(* Logix 5000 project; controller FV vendor 1 type 14 code 217 rev 31.11; software revision 31.00; part 14 of 63 *)
(* tags used below, declared in another part *)
   CWD : CHECKWORD_FLAGS;
   FR_B240 : INT[255];   // DEBOUNCE Debounce Flags
   FR_B246 : INT[255];   // V_REVERSE Flags for reversing contol action
   FR_B3 : INT[255];   // BINARY
   FR_data_file_value_to_move : DINT;
   FR_F102 : REAL[20];
   FR_FV31_AV01 : PlantItem;   // FV31_AV01
   FR_FV31_AV04 : PlantItem;   // FV31_AV04
   FR_FV31_AV05 : PlantItem;   // FV31_AV05
   FR_FV31_AV06 : PlantItem;   // FV31_AV06
   FR_FV31_AV07 : PlantItem;   // FV31_AV07
   FR_FV31_ROTO : PlantItem;   // FV31_ROTO
   FR_FV31_VA01 : PlantItem;   // FV31_VA01
   FR_N10 : INT[265];   // FV_AGING Comms to FV Aging PL C
   FR_N100 : INT[265];   // FV FILLING
   FR_N110 : INT[265];   // GREEN BEER Green Beer Main
   FR_N120 : INT[265];   // YEAST CROP Yeast Cropping Main
   FR_N13 : INT[265];   // MV_ROUTE Comms to MV Routing PLC
   FR_N130 : INT[265];   // FILTRATE Filtrate Return
   FR_N14 : INT[265];   // MVFV CIP Comms to MVFV CIP Un it PLC
   FR_N160 : INT[265];   // VESSEL Vessel Working Direc tory
   FR_N200 : INT[265];   // ANALOG_IN Analog Inputs
   FR_N255 : INT[265];   // CHECKWORDS
   FR_N31 : INT[265];   // FV31
   FR_N7 : INT[265];   // INTEGER
   FR_N99 : INT[265];   // COMMENT Comment Lines
   FR_OXY_SW1 : PlantItem;   // OXY_SW1
   FR_OXY_SW2 : PlantItem;   // OXY_SW2
   FR_T101 : TIMER[255];   // FV FILLING
   FR_T144 : TIMER[255];   // CIP
   FR_T4 : TIMER[255];   // TIMER
   FR_T50 : TIMER[52];
   FR_T51 : TIMER[52];
   FR_T52 : TIMER[52];
   FR_T53 : TIMER[52];
   FR_VB1_AV08 : PlantItem;   // VB1_AV08
   FR_VB1_AV09 : PlantItem;   // VB1_AV09
   FR_VB2_AV04 : PlantItem;   // VB2_AV04
   FR_VB2_AV05 : PlantItem;   // VB2_AV05
   FR_VB3_AV04 : PlantItem;   // VB3_AV04
   FR_VB3_AV05 : PlantItem;   // VB3_AV05
   FR_VB4_AV03 : PlantItem;   // VB4_AV03
   FR_VB4_AV09 : PlantItem;   // VB4_AV09
   FR_VB4_AV15 : PlantItem;   // VB4_AV15
(* FR_Common, continued *)

ROUTINE FR_FV31_31   (* ladder *)
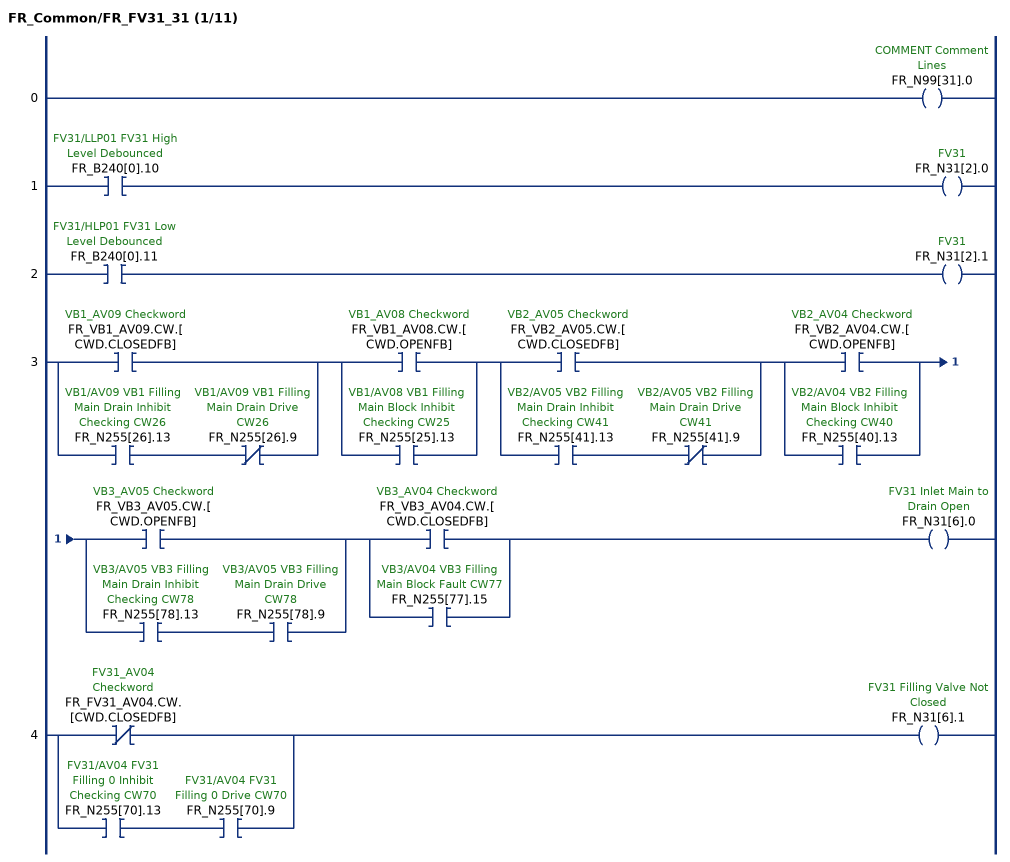
   0: OTE(FR_N99[31].0);
   1: XIC(FR_B240[0].10)OTE(FR_N31[2].0);
   2: XIC(FR_B240[0].11)OTE(FR_N31[2].1);
   3: [XIC(FR_VB1_AV09.CW.[CWD.CLOSEDFB]) ,XIC(FR_N255[26].13) XIO(FR_N255[26].9) ][XIC(FR_VB1_AV08.CW.[CWD.OPENFB]) ,XIC(FR_N255[25].13) ][XIC(FR_VB2_AV05.CW.[CWD.CLOSEDFB]) ,XIC(FR_N255[41].13) XIO(FR_N255[41].9) ][XIC(FR_VB2_AV04.CW.[CWD.OPENFB]) ,XIC(FR_N255[40].13) ][XIC(FR_VB3_AV05.CW.[CWD.OPENFB]) ,XIC(FR_N255[78].13) XIC(FR_N255[78].9) ][XIC(FR_VB3_AV04.CW.[CWD.CLOSEDFB]) ,XIC(FR_N255[77].15) ]OTE(FR_N31[6].0);
   4: [XIO(FR_FV31_AV04.CW.[CWD.CLOSEDFB]) ,XIC(FR_N255[70].13) XIC(FR_N255[70].9) ]OTE(FR_N31[6].1);
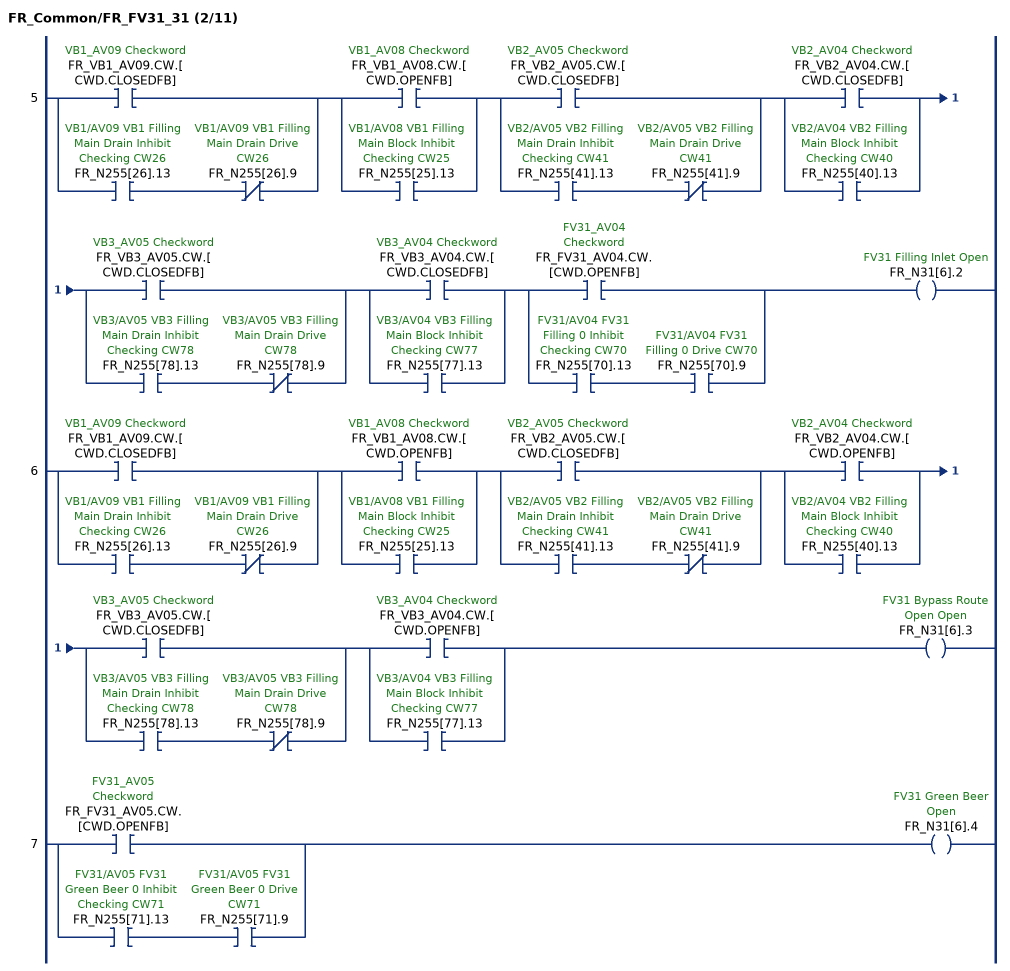
   5: [XIC(FR_VB1_AV09.CW.[CWD.CLOSEDFB]) ,XIC(FR_N255[26].13) XIO(FR_N255[26].9) ][XIC(FR_VB1_AV08.CW.[CWD.OPENFB]) ,XIC(FR_N255[25].13) ][XIC(FR_VB2_AV05.CW.[CWD.CLOSEDFB]) ,XIC(FR_N255[41].13) XIO(FR_N255[41].9) ][XIC(FR_VB2_AV04.CW.[CWD.CLOSEDFB]) ,XIC(FR_N255[40].13) ][XIC(FR_VB3_AV05.CW.[CWD.CLOSEDFB]) ,XIC(FR_N255[78].13) XIO(FR_N255[78].9) ][XIC(FR_VB3_AV04.CW.[CWD.CLOSEDFB]) ,XIC(FR_N255[77].13) ][XIC(FR_FV31_AV04.CW.[CWD.OPENFB]) ,XIC(FR_N255[70].13) XIC(FR_N255[70].9) ]OTE(FR_N31[6].2);
   6: [XIC(FR_VB1_AV09.CW.[CWD.CLOSEDFB]) ,XIC(FR_N255[26].13) XIO(FR_N255[26].9) ][XIC(FR_VB1_AV08.CW.[CWD.OPENFB]) ,XIC(FR_N255[25].13) ][XIC(FR_VB2_AV05.CW.[CWD.CLOSEDFB]) ,XIC(FR_N255[41].13) XIO(FR_N255[41].9) ][XIC(FR_VB2_AV04.CW.[CWD.OPENFB]) ,XIC(FR_N255[40].13) ][XIC(FR_VB3_AV05.CW.[CWD.CLOSEDFB]) ,XIC(FR_N255[78].13) XIO(FR_N255[78].9) ][XIC(FR_VB3_AV04.CW.[CWD.OPENFB]) ,XIC(FR_N255[77].13) ]OTE(FR_N31[6].3);
   7: [XIC(FR_FV31_AV05.CW.[CWD.OPENFB]) ,XIC(FR_N255[71].13) XIC(FR_N255[71].9) ]OTE(FR_N31[6].4);
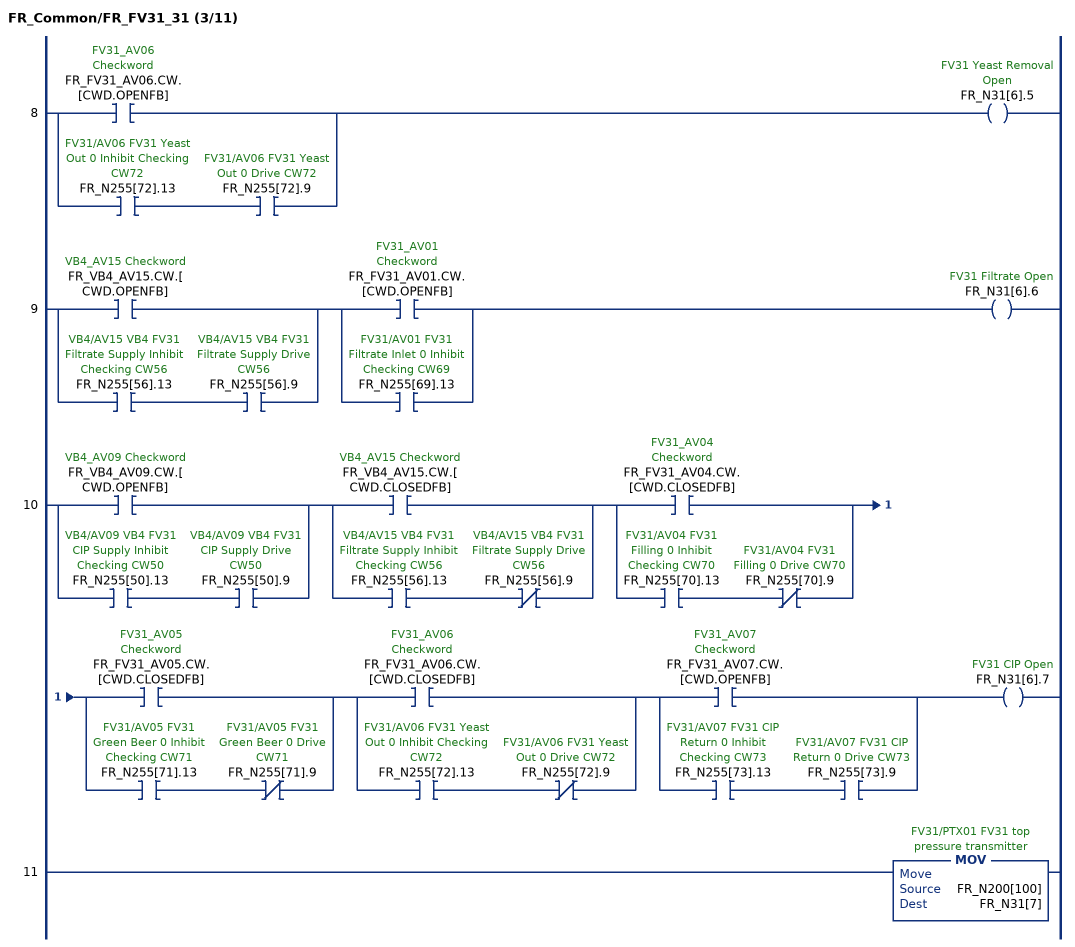
   8: [XIC(FR_FV31_AV06.CW.[CWD.OPENFB]) ,XIC(FR_N255[72].13) XIC(FR_N255[72].9) ]OTE(FR_N31[6].5);
   9: [XIC(FR_VB4_AV15.CW.[CWD.OPENFB]) ,XIC(FR_N255[56].13) XIC(FR_N255[56].9) ][XIC(FR_FV31_AV01.CW.[CWD.OPENFB]) ,XIC(FR_N255[69].13) ]OTE(FR_N31[6].6);
   10: [XIC(FR_VB4_AV09.CW.[CWD.OPENFB]) ,XIC(FR_N255[50].13) XIC(FR_N255[50].9) ][XIC(FR_VB4_AV15.CW.[CWD.CLOSEDFB]) ,XIC(FR_N255[56].13) XIO(FR_N255[56].9) ][XIC(FR_FV31_AV04.CW.[CWD.CLOSEDFB]) ,XIC(FR_N255[70].13) XIO(FR_N255[70].9) ][XIC(FR_FV31_AV05.CW.[CWD.CLOSEDFB]) ,XIC(FR_N255[71].13) XIO(FR_N255[71].9) ][XIC(FR_FV31_AV06.CW.[CWD.CLOSEDFB]) ,XIC(FR_N255[72].13) XIO(FR_N255[72].9) ][XIC(FR_FV31_AV07.CW.[CWD.OPENFB]) ,XIC(FR_N255[73].13) XIC(FR_N255[73].9) ]OTE(FR_N31[6].7);
   11: MOV(FR_N200[100],FR_N31[7]);
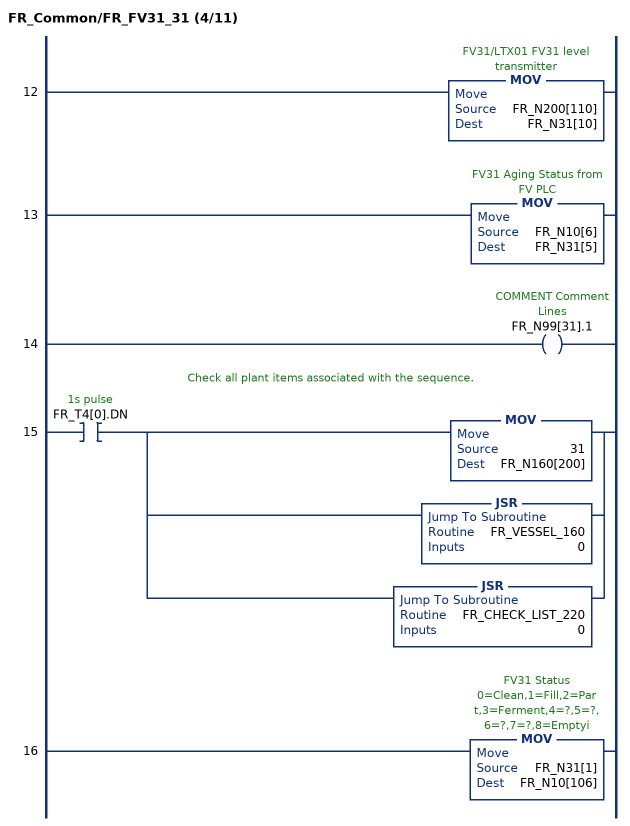
   12: MOV(FR_N200[110],FR_N31[10]);
   13: MOV(FR_N10[6],FR_N31[5]);
   14: OTE(FR_N99[31].1);
   // Check all plant items associated with the sequence.
   15: XIC(FR_T4[0].DN)[MOV(31,FR_N160[200]) ,JSR(FR_VESSEL_160,0) ,JSR(FR_CHECK_LIST_220,0) ];
   16: MOV(FR_N31[1],FR_N10[106]);
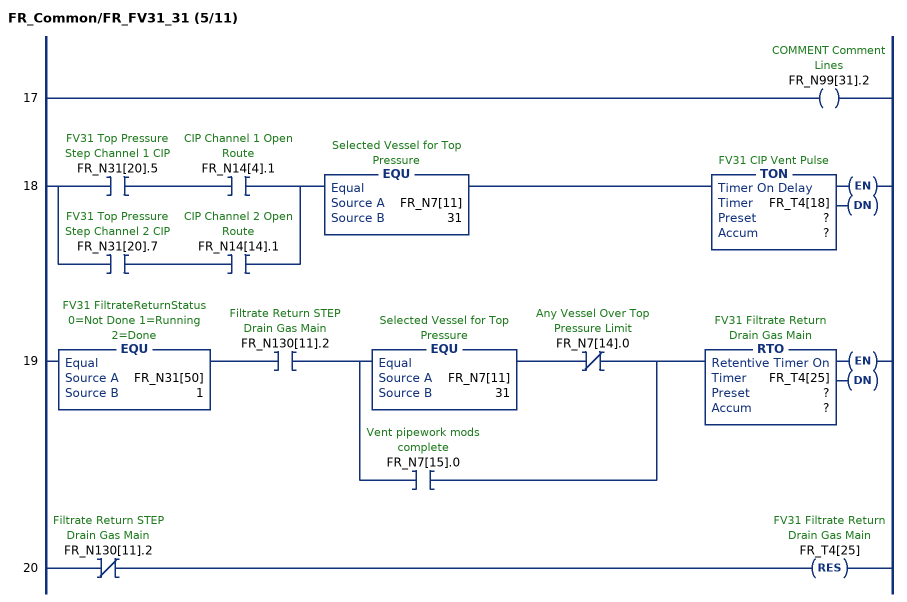
   17: OTE(FR_N99[31].2);
   18: [XIC(FR_N31[20].5) XIC(FR_N14[4].1) ,XIC(FR_N31[20].7) XIC(FR_N14[14].1) ]EQU(FR_N7[11],31)TON(FR_T4[18],?,?);
   19: EQU(FR_N31[50],1)XIC(FR_N130[11].2)[EQU(FR_N7[11],31) XIO(FR_N7[14].0) ,XIC(FR_N7[15].0) ]RTO(FR_T4[25],?,?);
   20: XIO(FR_N130[11].2)RES(FR_T4[25]);
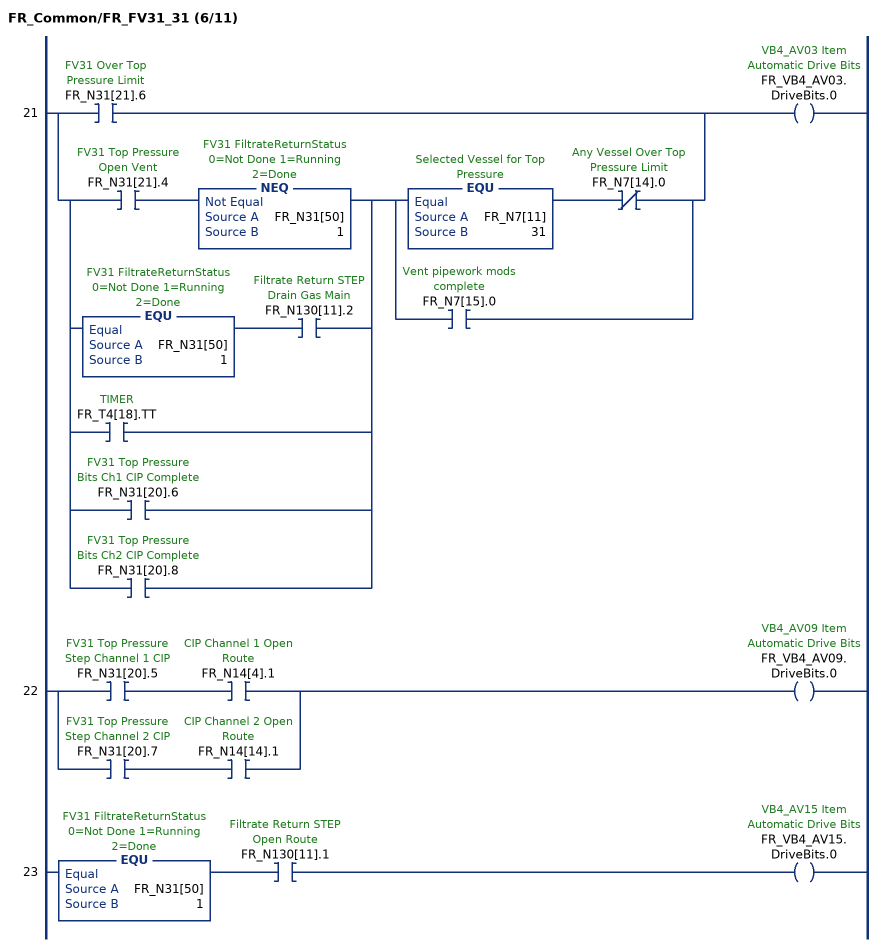
   21: [XIC(FR_N31[21].6) ,[XIC(FR_N31[21].4) NEQ(FR_N31[50],1) ,EQU(FR_N31[50],1) XIC(FR_N130[11].2) ,XIC(FR_T4[18].TT) ,[XIC(FR_N31[20].6) ,XIC(FR_N31[20].8) ] ] [EQU(FR_N7[11],31) XIO(FR_N7[14].0) ,XIC(FR_N7[15].0) ] ]OTE(FR_VB4_AV03.DriveBits.0);
   22: [XIC(FR_N31[20].5) XIC(FR_N14[4].1) ,XIC(FR_N31[20].7) XIC(FR_N14[14].1) ]OTE(FR_VB4_AV09.DriveBits.0);
   23: EQU(FR_N31[50],1)XIC(FR_N130[11].1)OTE(FR_VB4_AV15.DriveBits.0);
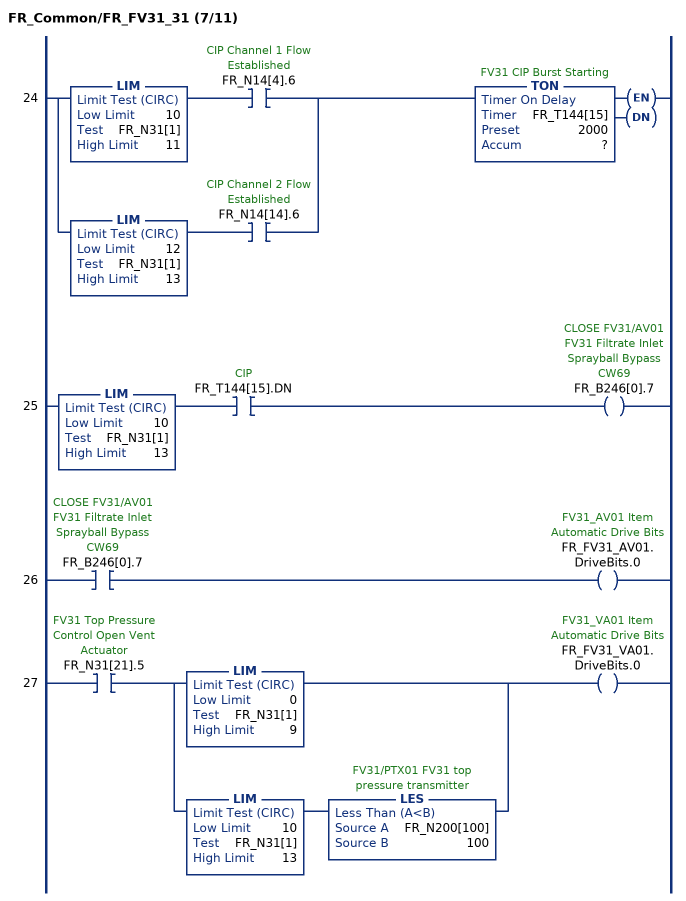
   24: [LIM(10,FR_N31[1],11) XIC(FR_N14[4].6) ,LIM(12,FR_N31[1],13) XIC(FR_N14[14].6) ]TON(FR_T144[15],?,?);
   25: LIM(10,FR_N31[1],13)XIC(FR_T144[15].DN)OTE(FR_B246[0].7);
   26: XIC(FR_B246[0].7)OTE(FR_FV31_AV01.DriveBits.0);
   27: XIC(FR_N31[21].5)[LIM(0,FR_N31[1],9) ,LIM(10,FR_N31[1],13) LES(FR_N200[100],100) ]OTE(FR_FV31_VA01.DriveBits.0);
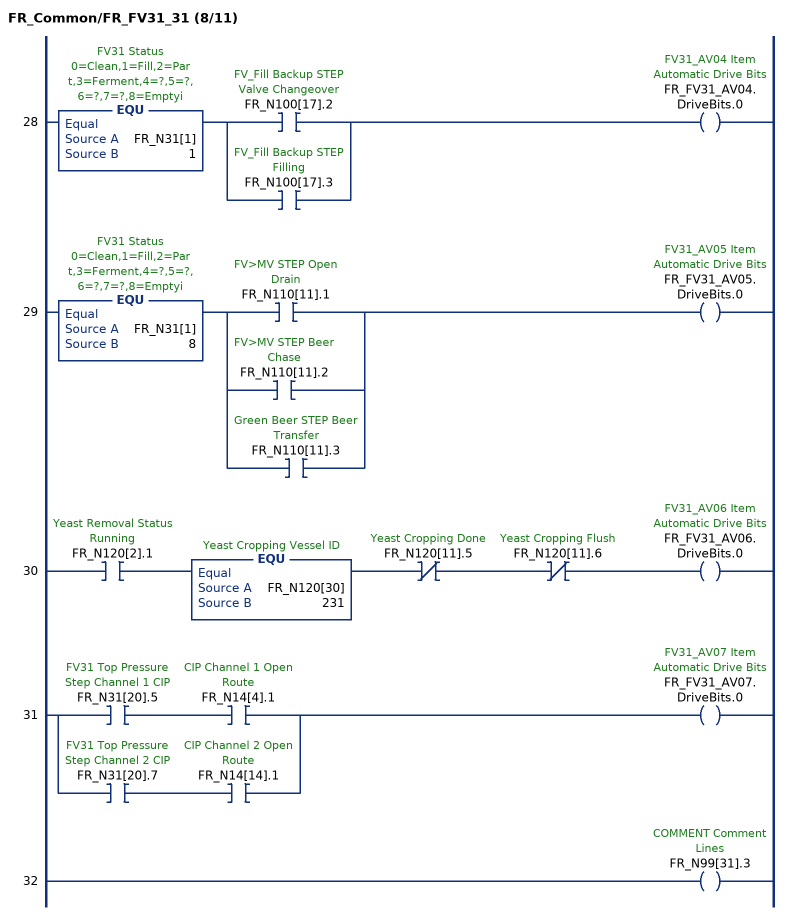
   28: EQU(FR_N31[1],1)[XIC(FR_N100[17].2) ,XIC(FR_N100[17].3) ]OTE(FR_FV31_AV04.DriveBits.0);
   29: EQU(FR_N31[1],8)[XIC(FR_N110[11].1) ,XIC(FR_N110[11].2) ,XIC(FR_N110[11].3) ]OTE(FR_FV31_AV05.DriveBits.0);
   30: XIC(FR_N120[2].1)EQU(FR_N120[30],231)XIO(FR_N120[11].5)XIO(FR_N120[11].6)OTE(FR_FV31_AV06.DriveBits.0);
   31: [XIC(FR_N31[20].5) XIC(FR_N14[4].1) ,XIC(FR_N31[20].7) XIC(FR_N14[14].1) ]OTE(FR_FV31_AV07.DriveBits.0);
   32: OTE(FR_N99[31].3);
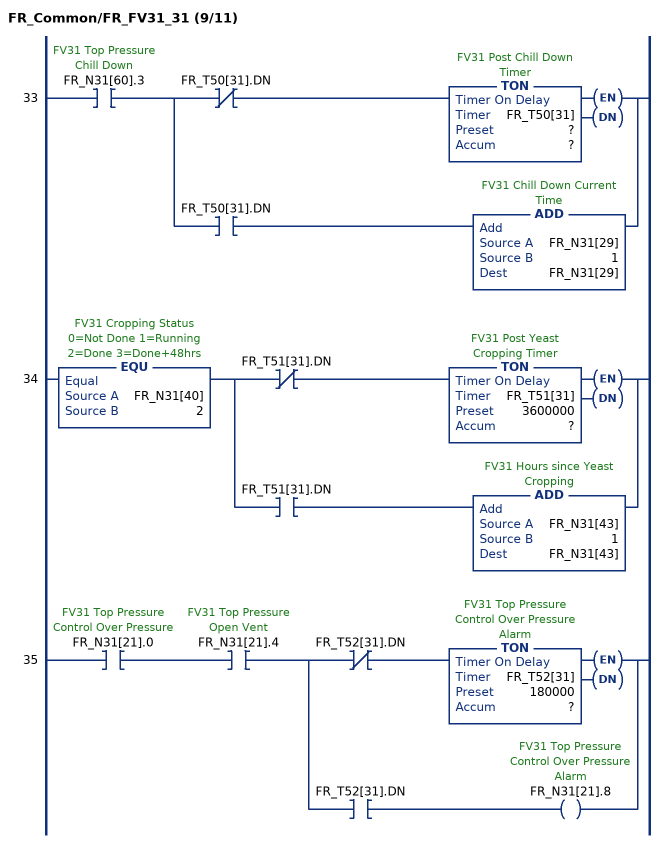
   33: XIC(FR_N31[60].3)[XIO(FR_T50[31].DN) TON(FR_T50[31],?,?) ,XIC(FR_T50[31].DN) ADD(FR_N31[29],1,FR_N31[29]) ];
   34: EQU(FR_N31[40],2)[XIO(FR_T51[31].DN) TON(FR_T51[31],?,?) ,XIC(FR_T51[31].DN) ADD(FR_N31[43],1,FR_N31[43]) ];
   35: XIC(FR_N31[21].0)XIC(FR_N31[21].4)[XIO(FR_T52[31].DN) TON(FR_T52[31],?,?) ,XIC(FR_T52[31].DN) OTE(FR_N31[21].8) ];
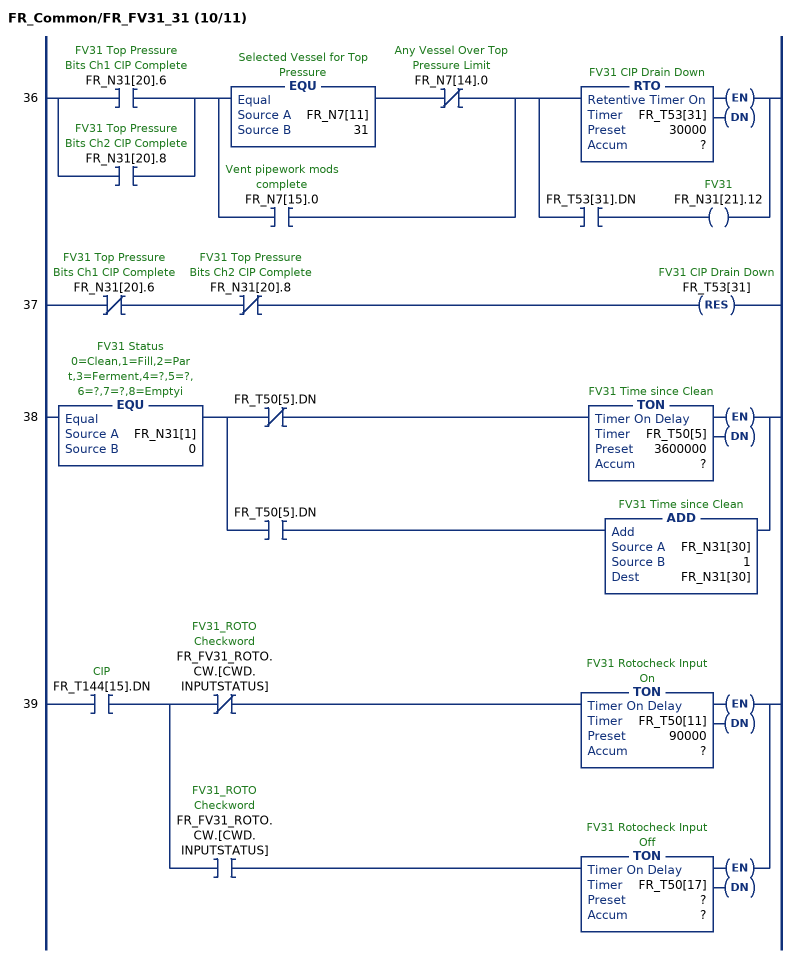
   36: [XIC(FR_N31[20].6) ,XIC(FR_N31[20].8) ][EQU(FR_N7[11],31) XIO(FR_N7[14].0) ,XIC(FR_N7[15].0) ][RTO(FR_T53[31],?,?) ,XIC(FR_T53[31].DN) OTE(FR_N31[21].12) ];
   37: XIO(FR_N31[20].6)XIO(FR_N31[20].8)RES(FR_T53[31]);
   38: EQU(FR_N31[1],0)[XIO(FR_T50[5].DN) TON(FR_T50[5],?,?) ,XIC(FR_T50[5].DN) ADD(FR_N31[30],1,FR_N31[30]) ];
   39: XIC(FR_T144[15].DN)[XIO(FR_FV31_ROTO.CW.[CWD.INPUTSTATUS]) TON(FR_T50[11],?,?) ,XIC(FR_FV31_ROTO.CW.[CWD.INPUTSTATUS]) TON(FR_T50[17],?,?) ];
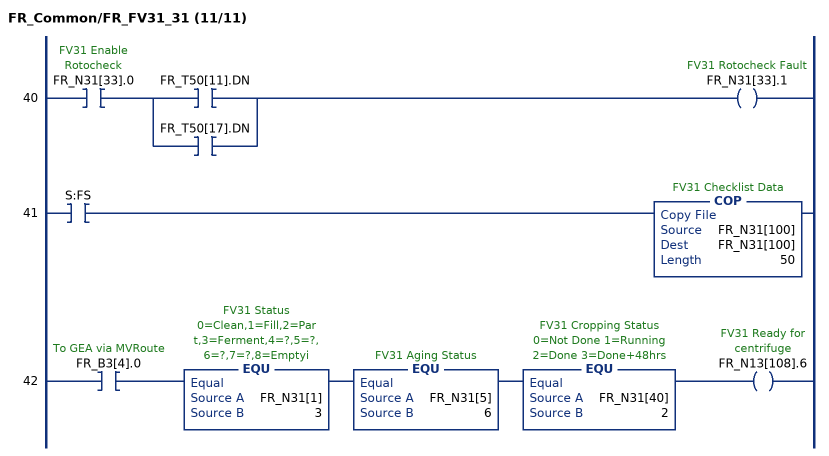
   40: XIC(FR_N31[33].0)[XIC(FR_T50[11].DN) ,XIC(FR_T50[17].DN) ]OTE(FR_N31[33].1);
   41: XIC(S:FS)COP(FR_N31[100],FR_N31[100],50);
   42: XIC(FR_B3[4].0)EQU(FR_N31[1],3)EQU(FR_N31[5],6)EQU(FR_N31[40],2)OTE(FR_N13[108].6);
END_ROUTINE

ROUTINE FR_FV_FILL_101   (* ladder *)
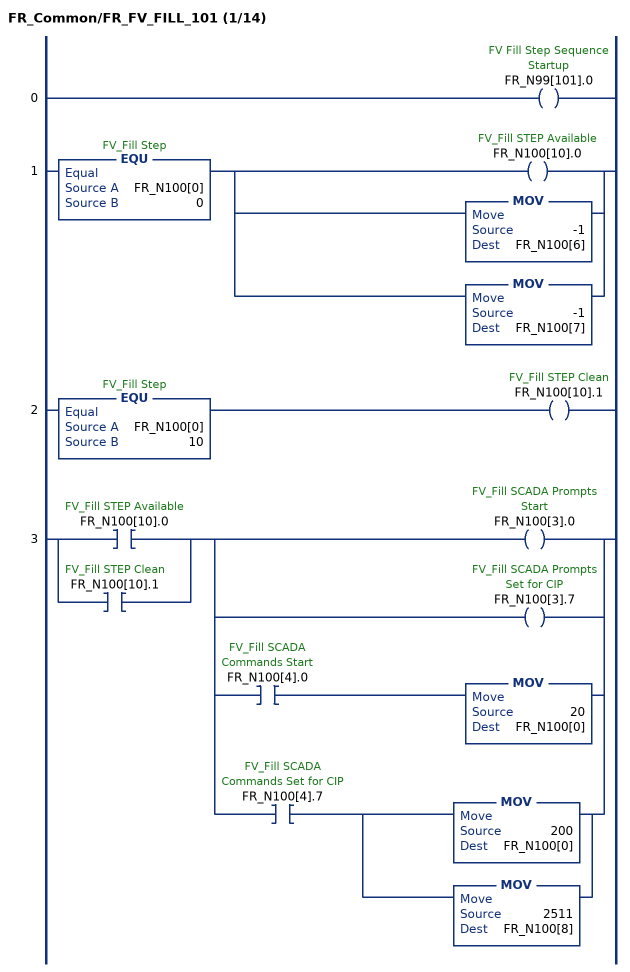
   0: OTE(FR_N99[101].0);
   1: EQU(FR_N100[0],0)[OTE(FR_N100[10].0) ,MOV(-1,FR_N100[6]) ,MOV(-1,FR_N100[7]) ];
   2: EQU(FR_N100[0],10)OTE(FR_N100[10].1);
   3: [XIC(FR_N100[10].0) ,XIC(FR_N100[10].1) ][OTE(FR_N100[3].0) ,OTE(FR_N100[3].7) ,XIC(FR_N100[4].0) MOV(20,FR_N100[0]) ,XIC(FR_N100[4].7) [MOV(200,FR_N100[0]) ,MOV(2511,FR_N100[8]) ] ];
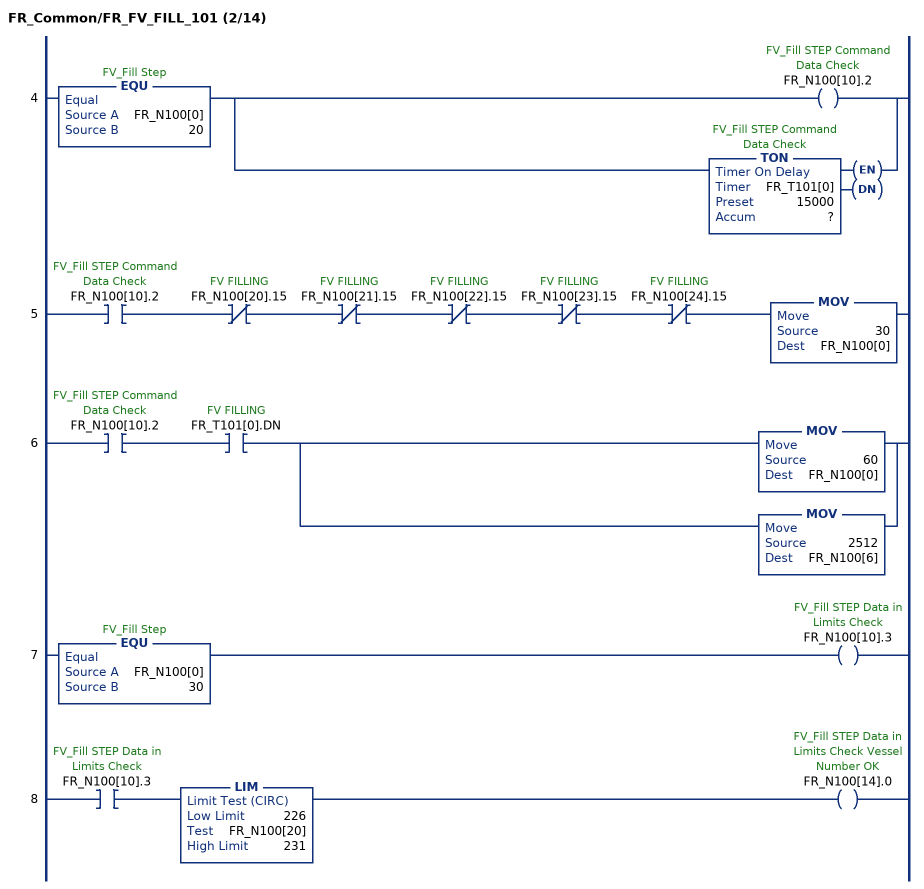
   4: EQU(FR_N100[0],20)[OTE(FR_N100[10].2) ,TON(FR_T101[0],?,?) ];
   5: XIC(FR_N100[10].2)XIO(FR_N100[20].15)XIO(FR_N100[21].15)XIO(FR_N100[22].15)XIO(FR_N100[23].15)XIO(FR_N100[24].15)MOV(30,FR_N100[0]);
   6: XIC(FR_N100[10].2)XIC(FR_T101[0].DN)[MOV(60,FR_N100[0]) ,MOV(2512,FR_N100[6]) ];
   7: EQU(FR_N100[0],30)OTE(FR_N100[10].3);
   8: XIC(FR_N100[10].3)LIM(226,FR_N100[20],231)OTE(FR_N100[14].0);
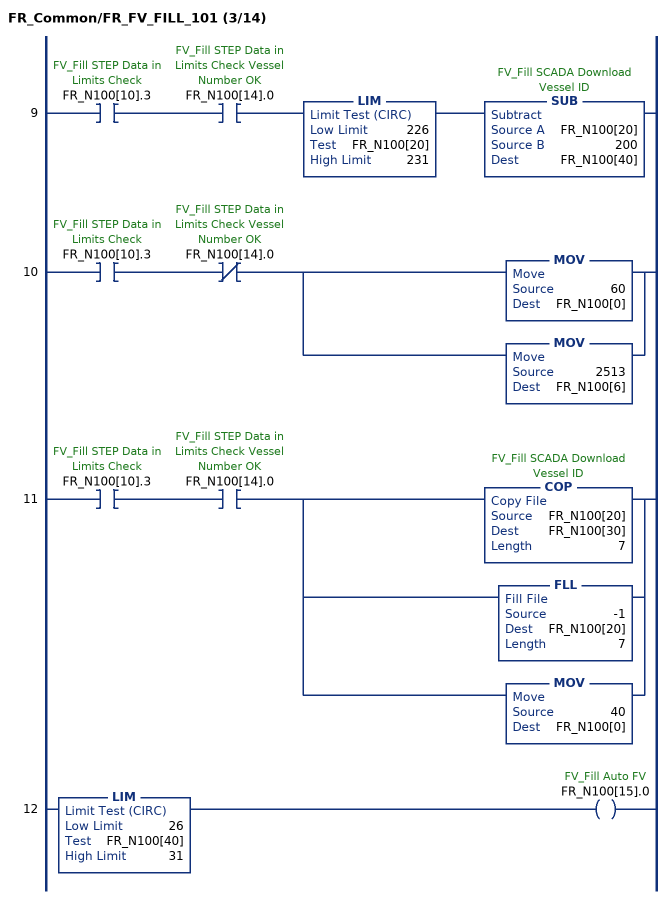
   9: XIC(FR_N100[10].3)XIC(FR_N100[14].0)LIM(226,FR_N100[20],231)SUB(FR_N100[20],200,FR_N100[40]);
   10: XIC(FR_N100[10].3)XIO(FR_N100[14].0)[MOV(60,FR_N100[0]) ,MOV(2513,FR_N100[6]) ];
   11: XIC(FR_N100[10].3)XIC(FR_N100[14].0)[COP(FR_N100[20],FR_N100[30],7) ,FLL(-1,FR_N100[20],7) ,MOV(40,FR_N100[0]) ];
   12: LIM(26,FR_N100[40],31)OTE(FR_N100[15].0);
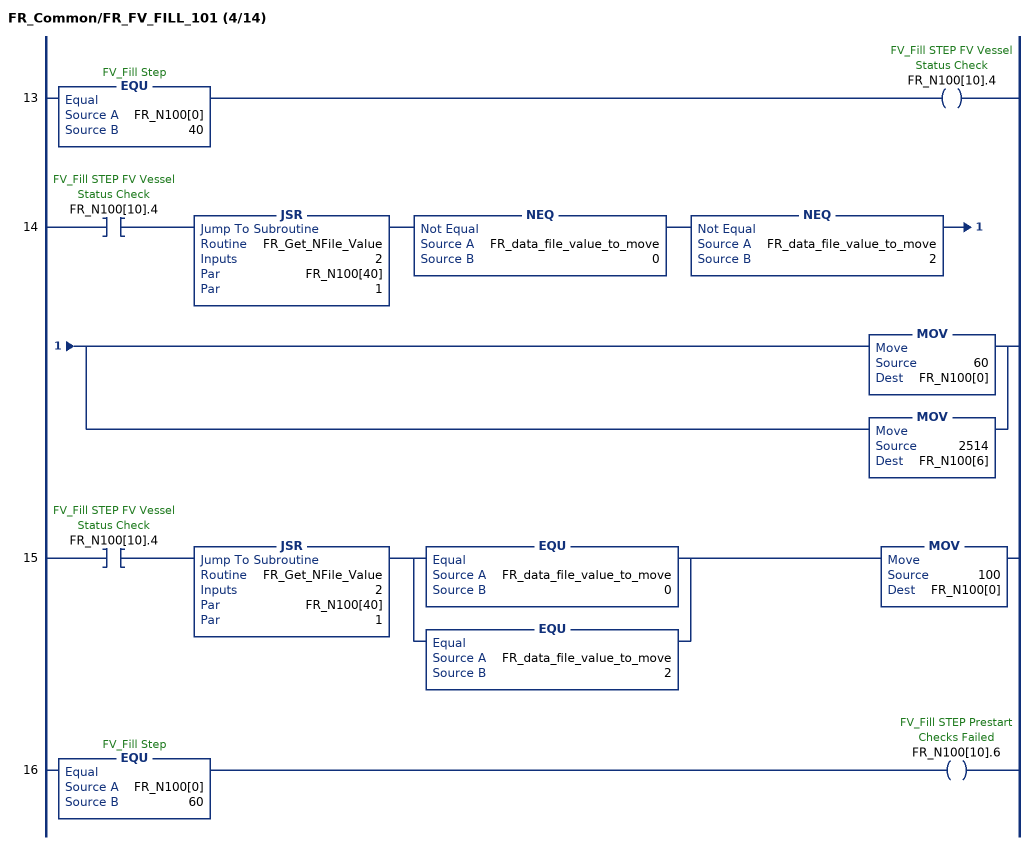
   13: EQU(FR_N100[0],40)OTE(FR_N100[10].4);
   14: XIC(FR_N100[10].4)JSR(FR_Get_NFile_Value,2,FR_N100[40],1)NEQ(FR_data_file_value_to_move,0)NEQ(FR_data_file_value_to_move,2)[MOV(60,FR_N100[0]) ,MOV(2514,FR_N100[6]) ];
   15: XIC(FR_N100[10].4)JSR(FR_Get_NFile_Value,2,FR_N100[40],1)[EQU(FR_data_file_value_to_move,0) ,EQU(FR_data_file_value_to_move,2) ]MOV(100,FR_N100[0]);
   16: EQU(FR_N100[0],60)OTE(FR_N100[10].6);
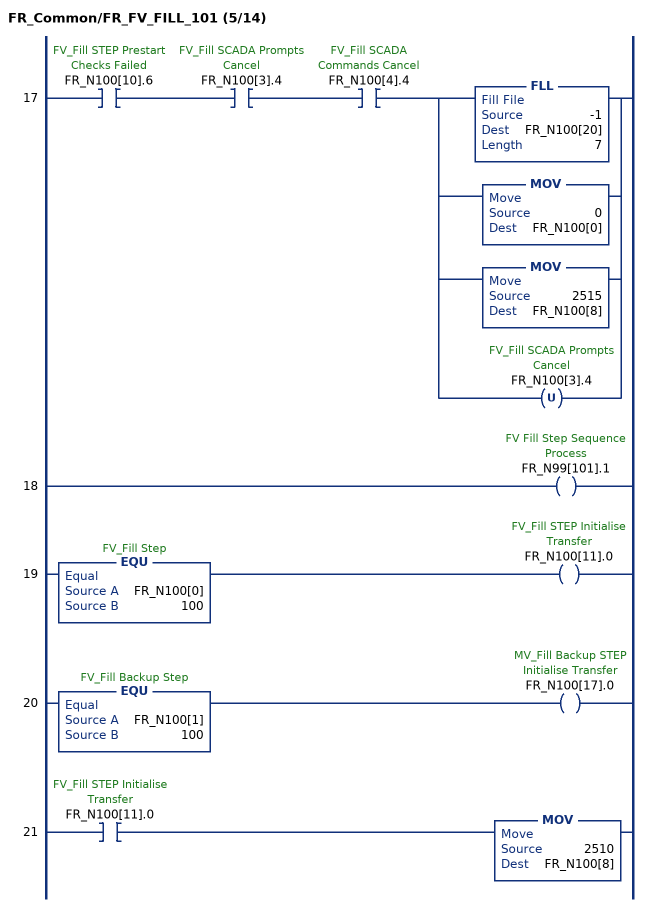
   17: XIC(FR_N100[10].6)XIC(FR_N100[3].4)XIC(FR_N100[4].4)[FLL(-1,FR_N100[20],7) ,MOV(0,FR_N100[0]) ,MOV(2515,FR_N100[8]) ,OTU(FR_N100[3].4) ];
   18: OTE(FR_N99[101].1);
   19: EQU(FR_N100[0],100)OTE(FR_N100[11].0);
   20: EQU(FR_N100[1],100)OTE(FR_N100[17].0);
   21: XIC(FR_N100[11].0)MOV(2510,FR_N100[8]);
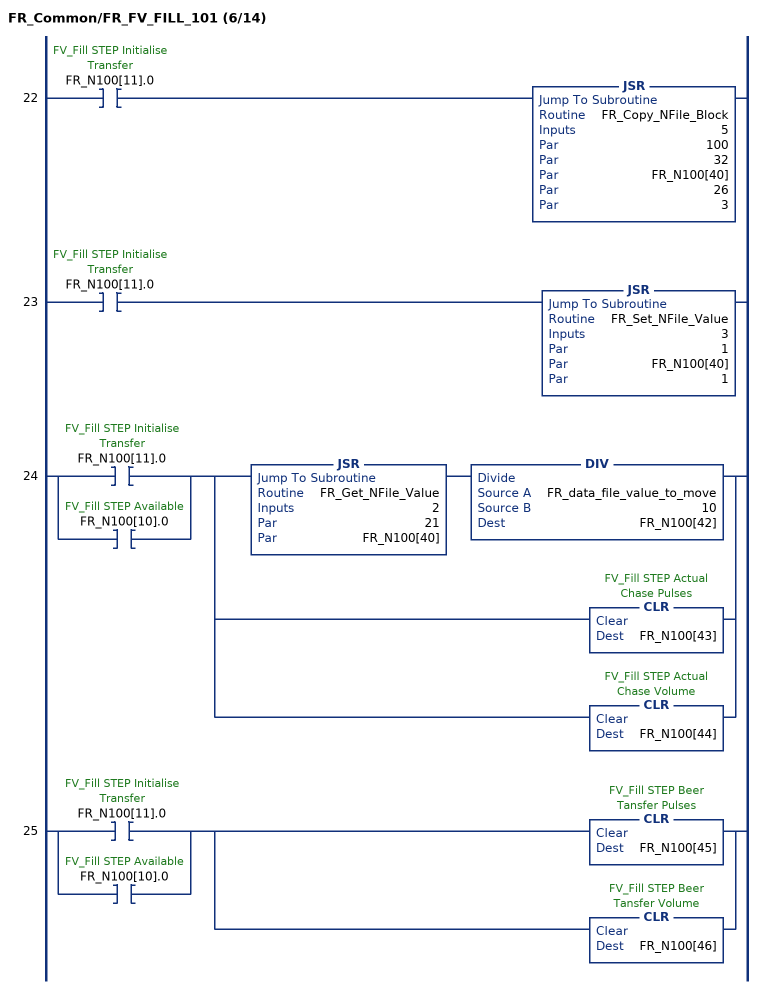
   22: XIC(FR_N100[11].0)JSR(FR_Copy_NFile_Block,5,100,32,FR_N100[40],26,3);
   23: XIC(FR_N100[11].0)JSR(FR_Set_NFile_Value,3,1,FR_N100[40],1);
   24: [XIC(FR_N100[11].0) ,XIC(FR_N100[10].0) ][JSR(FR_Get_NFile_Value,2,21,FR_N100[40]) DIV(FR_data_file_value_to_move,10,FR_N100[42]) ,CLR(FR_N100[43]) ,CLR(FR_N100[44]) ];
   25: [XIC(FR_N100[11].0) ,XIC(FR_N100[10].0) ][CLR(FR_N100[45]) ,CLR(FR_N100[46]) ];
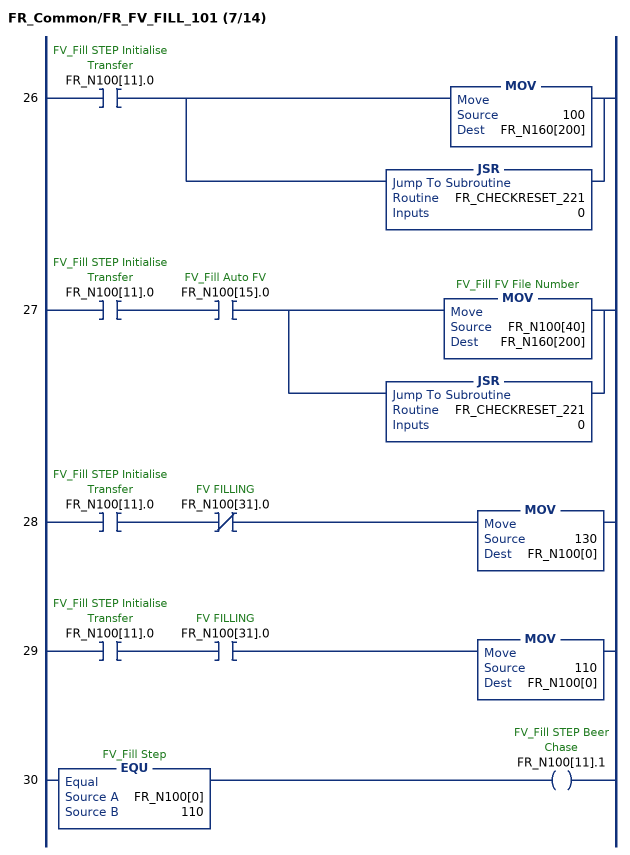
   26: XIC(FR_N100[11].0)[MOV(100,FR_N160[200]) ,JSR(FR_CHECKRESET_221,0) ];
   27: XIC(FR_N100[11].0)XIC(FR_N100[15].0)[MOV(FR_N100[40],FR_N160[200]) ,JSR(FR_CHECKRESET_221,0) ];
   28: XIC(FR_N100[11].0)XIO(FR_N100[31].0)MOV(130,FR_N100[0]);
   29: XIC(FR_N100[11].0)XIC(FR_N100[31].0)MOV(110,FR_N100[0]);
   30: EQU(FR_N100[0],110)OTE(FR_N100[11].1);
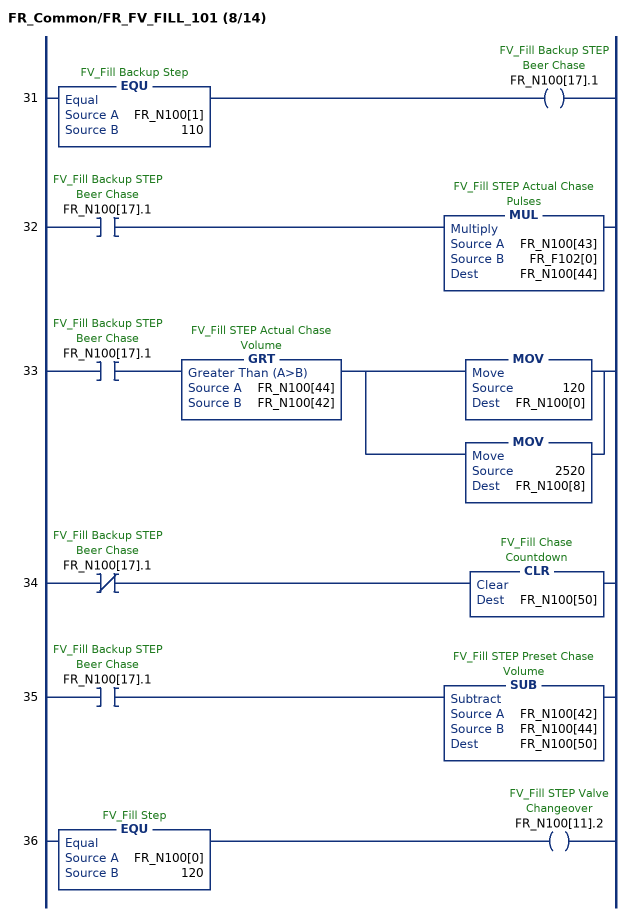
   31: EQU(FR_N100[1],110)OTE(FR_N100[17].1);
   32: XIC(FR_N100[17].1)MUL(FR_N100[43],FR_F102[0],FR_N100[44]);
   33: XIC(FR_N100[17].1)GRT(FR_N100[44],FR_N100[42])[MOV(120,FR_N100[0]) ,MOV(2520,FR_N100[8]) ];
   34: XIO(FR_N100[17].1)CLR(FR_N100[50]);
   35: XIC(FR_N100[17].1)SUB(FR_N100[42],FR_N100[44],FR_N100[50]);
   36: EQU(FR_N100[0],120)OTE(FR_N100[11].2);
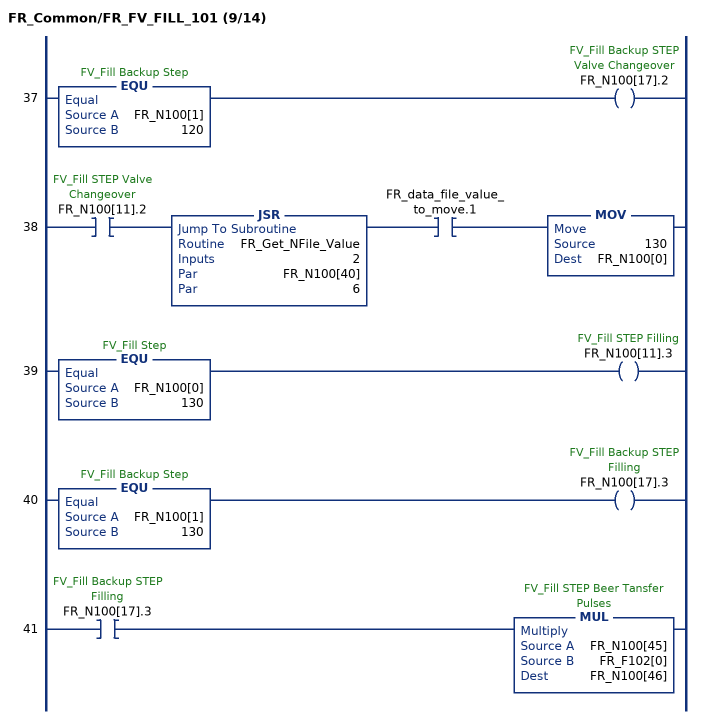
   37: EQU(FR_N100[1],120)OTE(FR_N100[17].2);
   38: XIC(FR_N100[11].2)JSR(FR_Get_NFile_Value,2,FR_N100[40],6)XIC(FR_data_file_value_to_move.1)MOV(130,FR_N100[0]);
   39: EQU(FR_N100[0],130)OTE(FR_N100[11].3);
   40: EQU(FR_N100[1],130)OTE(FR_N100[17].3);
   41: XIC(FR_N100[17].3)MUL(FR_N100[45],FR_F102[0],FR_N100[46]);
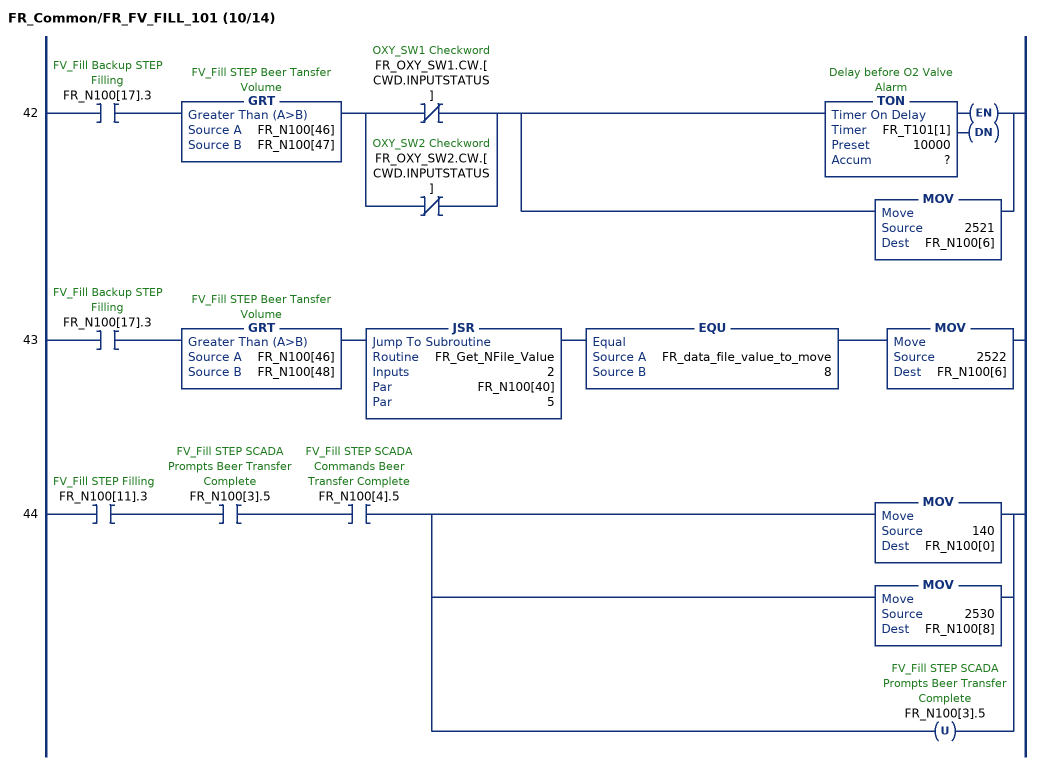
   42: XIC(FR_N100[17].3)GRT(FR_N100[46],FR_N100[47])[XIO(FR_OXY_SW1.CW.[CWD.INPUTSTATUS]) ,XIO(FR_OXY_SW2.CW.[CWD.INPUTSTATUS]) ][TON(FR_T101[1],?,?) ,MOV(2521,FR_N100[6]) ];
   43: XIC(FR_N100[17].3)GRT(FR_N100[46],FR_N100[48])JSR(FR_Get_NFile_Value,2,FR_N100[40],5)EQU(FR_data_file_value_to_move,8)MOV(2522,FR_N100[6]);
   44: XIC(FR_N100[11].3)XIC(FR_N100[3].5)XIC(FR_N100[4].5)[MOV(140,FR_N100[0]) ,MOV(2530,FR_N100[8]) ,OTU(FR_N100[3].5) ];
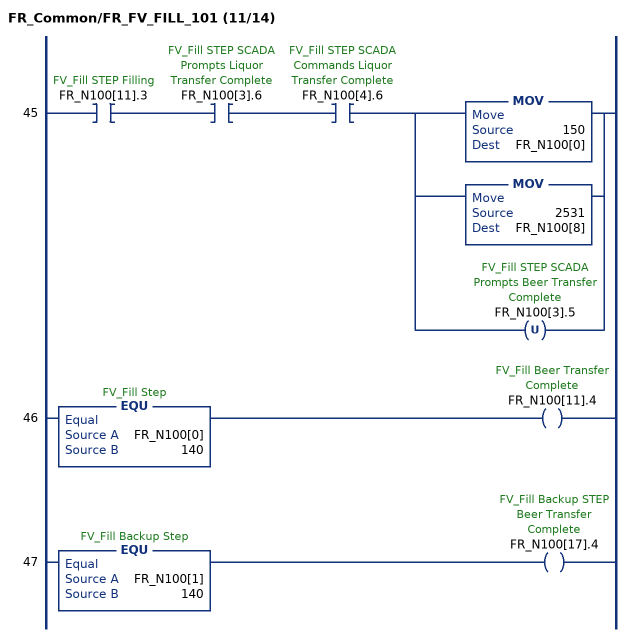
   45: XIC(FR_N100[11].3)XIC(FR_N100[3].6)XIC(FR_N100[4].6)[MOV(150,FR_N100[0]) ,MOV(2531,FR_N100[8]) ,OTU(FR_N100[3].5) ];
   46: EQU(FR_N100[0],140)OTE(FR_N100[11].4);
   47: EQU(FR_N100[1],140)OTE(FR_N100[17].4);
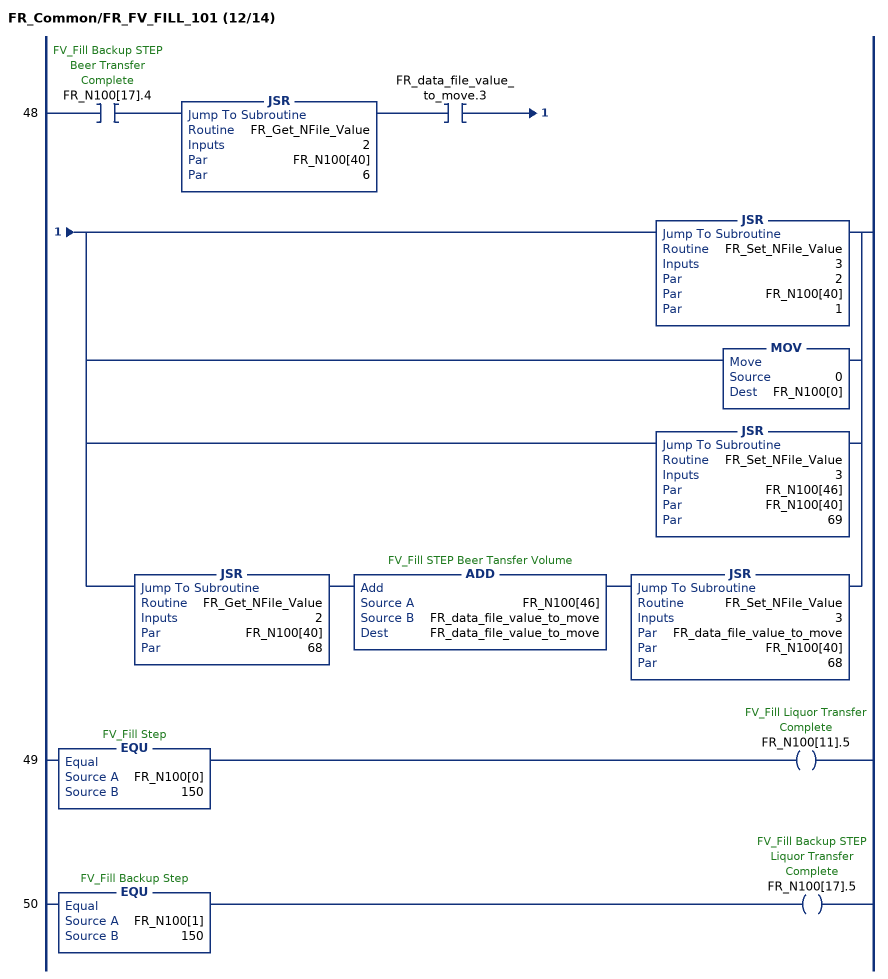
   48: XIC(FR_N100[17].4)JSR(FR_Get_NFile_Value,2,FR_N100[40],6)XIC(FR_data_file_value_to_move.3)[JSR(FR_Set_NFile_Value,3,2,FR_N100[40],1) ,MOV(0,FR_N100[0]) ,JSR(FR_Set_NFile_Value,3,FR_N100[46],FR_N100[40],69) ,JSR(FR_Get_NFile_Value,2,FR_N100[40],68) ADD(FR_N100[46],FR_data_file_value_to_move,FR_data_file_value_to_move) JSR(FR_Set_NFile_Value,3,FR_data_file_value_to_move,FR_N100[40],68) ];
   49: EQU(FR_N100[0],150)OTE(FR_N100[11].5);
   50: EQU(FR_N100[1],150)OTE(FR_N100[17].5);
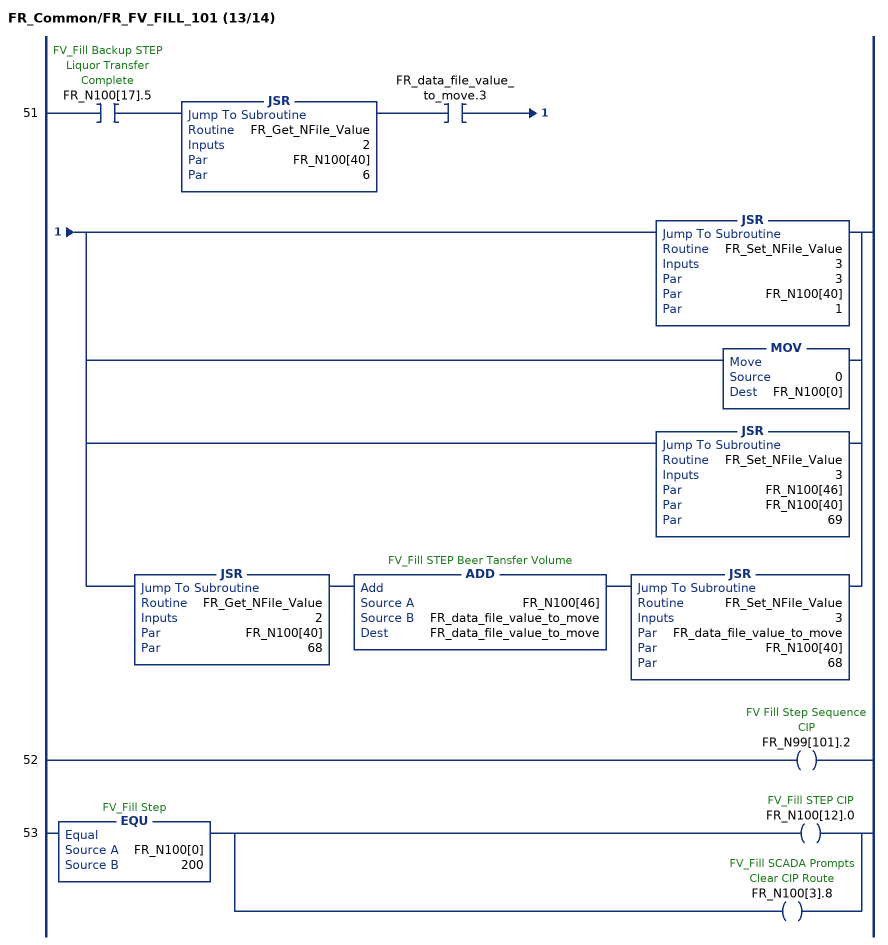
   51: XIC(FR_N100[17].5)JSR(FR_Get_NFile_Value,2,FR_N100[40],6)XIC(FR_data_file_value_to_move.3)[JSR(FR_Set_NFile_Value,3,3,FR_N100[40],1) ,MOV(0,FR_N100[0]) ,JSR(FR_Set_NFile_Value,3,FR_N100[46],FR_N100[40],69) ,JSR(FR_Get_NFile_Value,2,FR_N100[40],68) ADD(FR_N100[46],FR_data_file_value_to_move,FR_data_file_value_to_move) JSR(FR_Set_NFile_Value,3,FR_data_file_value_to_move,FR_N100[40],68) ];
   52: OTE(FR_N99[101].2);
   53: EQU(FR_N100[0],200)[OTE(FR_N100[12].0) ,OTE(FR_N100[3].8) ];
